
screen "MTA-ChillersBombasEnvasado" 800x480, template "Plantilla_2"
   GraphicView "Visor de gráficos_3" at 648,158 size 48x71; Picture "Bomba"
   GraphicIOField "Plantilla_Campo ES gráfico_2" at 684,217 size 49x36; PictureList "Motor2"
      ProcessValue <- "AnimaciónMT009"
   SymbolicIOField "Campo ES simbólico_4" at 602,132 size 172x21; TextOff '0'; TextOn '1'; TextList "EstadoMotor"
      ProcessValue <- "AnimaciónMT009"
   TextField "Campo de texto_6" at 599,93 size 42x18; Text 'MT009'
   GraphicView "Visor de gráficos_4" at 454,158 size 48x71; Picture "Bomba"
   GraphicIOField "Plantilla_Campo ES gráfico_1" at 490,217 size 49x36; PictureList "Motor2"
      ProcessValue <- "AnimaciónMT010"
   SymbolicIOField "Campo ES simbólico_1" at 408,132 size 172x21; TextOff '0'; TextOn '1'; TextList "EstadoMotor"
      ProcessValue <- "AnimaciónMT010"
   TextField "Campo de texto_7" at 405,93 size 42x18; Text 'MT010'
   GraphicView "Visor de gráficos_6" at 64,158 size 48x71; Picture "Bomba"
   GraphicIOField "Plantilla_Campo ES gráfico_4" at 100,217 size 49x36; PictureList "Motor2"
      ProcessValue <- "AnimaciónMP013"
   SymbolicIOField "Campo ES simbólico_3" at 20,132 size 172x21; TextOff '0'; TextOn '1'; TextList "EstadoMotor"
      ProcessValue <- "AnimaciónMP013"
   TextField "Campo de texto_9" at 23,93 size 41x18; Text 'MP013'
   TextField "Campo de texto_19" at 405,112 size 169x18; Text 'Intercambiador Línea 1 y Man.'
   GraphicView "Visor de gráficos_5" at 260,158 size 48x71; Picture "Bomba"
   GraphicIOField "Plantilla_Campo ES gráfico_3" at 296,217 size 49x36; PictureList "Motor2"
      ProcessValue <- "AnimaciónMP012"
   SymbolicIOField "Campo ES simbólico_2" at 214,132 size 172x21; TextOff '0'; TextOn '1'; TextList "EstadoMotor"
      ProcessValue <- "AnimaciónMP012"
   TextField "Campo de texto_8" at 211,93 size 41x18; Text 'MP012'
   TextField "Campo de texto_18" at 598,112 size 150x18; Text 'Intercambiador Línea 3 y 5'
   TextField "Campo de texto_16" at 215,113 size 150x18; Text 'Chillers Envasado - Principal'
   TextField "Campo de texto_17" at 21,113 size 146x18; Text 'Chillers Envasado - Backup'
   GraphicView "Plantilla_Visor de gráficos_2" at 752,6 size 35x35; Picture "ParlantesGris_1"
   GraphicView "Plantilla_Visor de gráficos_1" at 752,6 size 35x35; Picture "ParlantesRojo"
      Visibility <- "SirenaChillers"
   Button "Botón_1" at 740,1 size 57x44; TextOff 'Text'
      on Click: ActivateScreen("MTA-ChillersConfiguraciónSirena", 0)
   ScreenModuleView "ControlMotor-NoAUTO_1" at 609,271 size 163x76
      Guid_{11997190-67152} <- "DesMT009"
      Guid_{11997190-67156} <- "ParadaMT009"
      Guid_{11997190-67150} <- "HabMT009"
      Guid_{11997190-67154} <- "MarchaMT009"
   ScreenModuleView "ControlMotor-NoAUTO_2" at 413,271 size 163x76
      Guid_{11997190-67152} <- "DesMT010"
      Guid_{11997190-67156} <- "ParadaMT010"
      Guid_{11997190-67150} <- "HabMT010"
      Guid_{11997190-67154} <- "MarchaMT010"
   ScreenModuleView "ControlMotor-NoAUTO_3" at 219,271 size 163x76
      Guid_{11997190-67152} <- "DesMP012"
      Guid_{11997190-67156} <- "ParadaMP012"
      Guid_{11997190-67150} <- "HabMP012"
      Guid_{11997190-67154} <- "MarchaMP012"
   ScreenModuleView "ControlMotor-NoAUTO_4" at 22,271 size 163x76
      Guid_{11997190-67152} <- "DesMP013"
      Guid_{11997190-67156} <- "ParadaMP013"
      Guid_{11997190-67150} <- "HabMP013"
      Guid_{11997190-67154} <- "MarchaMP013"
   TextField "Campo de texto_5" at 256,10 size 261x27; Text 'Chillers - Bombas de Envasado'

screen "MTA-ChillersBombasSoplado" 800x480, template "Plantilla_2"
   TextField "Campo de texto_5" at 256,10 size 248x27; Text 'Chillers - Bombas de Soplado'
   GraphicView "Visor de gráficos_3" at 648,158 size 48x71; Picture "Bomba"
   GraphicIOField "Plantilla_Campo ES gráfico_8" at 684,217 size 49x36; PictureList "Motor2"
      ProcessValue <- "AnimaciónMT007"
   SymbolicIOField "Campo ES simbólico_4" at 602,132 size 172x21; TextOff '0'; TextOn '1'; TextList "EstadoMotor"
      ProcessValue <- "AnimaciónMT007"
   TextField "Campo de texto_6" at 599,93 size 42x18; Text 'MT007'
   GraphicView "Visor de gráficos_4" at 454,158 size 48x71; Picture "Bomba"
   GraphicIOField "Plantilla_Campo ES gráfico_7" at 490,217 size 49x36; PictureList "Motor2"
      ProcessValue <- "AnimaciónMT008"
   SymbolicIOField "Campo ES simbólico_1" at 408,132 size 172x21; TextOff '0'; TextOn '1'; TextList "EstadoMotor"
      ProcessValue <- "AnimaciónMT008"
   TextField "Campo de texto_7" at 405,93 size 42x18; Text 'MT008'
   GraphicView "Visor de gráficos_6" at 64,158 size 48x71; Picture "Bomba"
   GraphicIOField "Plantilla_Campo ES gráfico_5" at 100,217 size 49x36; PictureList "Motor2"
      ProcessValue <- "AnimaciónMP011"
   SymbolicIOField "Campo ES simbólico_3" at 20,132 size 172x21; TextOff '0'; TextOn '1'; TextList "EstadoMotor"
      ProcessValue <- "AnimaciónMP011"
   TextField "Campo de texto_9" at 23,93 size 41x18; Text 'MP011'
   TextField "Campo de texto_19" at 407,113 size 140x18; Text 'Sopladora Línea 3 y Man.'
   GraphicView "Visor de gráficos_5" at 260,158 size 48x71; Picture "Bomba"
   GraphicIOField "Plantilla_Campo ES gráfico_6" at 296,217 size 49x36; PictureList "Motor2"
      ProcessValue <- "AnimaciónMP010"
   SymbolicIOField "Campo ES simbólico_2" at 214,132 size 172x21; TextOff '0'; TextOn '1'; TextList "EstadoMotor"
      ProcessValue <- "AnimaciónMP010"
   TextField "Campo de texto_8" at 211,93 size 41x18; Text 'MP010'
   TextField "Campo de texto_18" at 599,113 size 104x18; Text 'Sopladora Línea 1'
   TextField "Campo de texto_16" at 212,113 size 142x18; Text 'Chillers Soplado - Principal'
   TextField "Campo de texto_17" at 21,113 size 138x18; Text 'Chillers Soplado - Backup'
   GraphicView "Plantilla_Visor de gráficos_2" at 752,6 size 35x35; Picture "ParlantesGris_1"
   GraphicView "Plantilla_Visor de gráficos_1" at 752,6 size 35x35; Picture "ParlantesRojo"
      Visibility <- "SirenaChillers"
   Button "Botón_1" at 740,1 size 57x44; TextOff 'Text'
      on Click: ActivateScreen("MTA-ChillersConfiguraciónSirena", 0)
   ScreenModuleView "ControlMotor-NoAUTO_1" at 609,271 size 163x76
      Guid_{11997190-67152} <- "DesMT007"
      Guid_{11997190-67156} <- "ParadaMT007"
      Guid_{11997190-67150} <- "HabMT007"
      Guid_{11997190-67154} <- "MarchaMT007"
   ScreenModuleView "ControlMotor-NoAUTO_3" at 219,271 size 163x76
      Guid_{11997190-67152} <- "DesMP010"
      Guid_{11997190-67156} <- "ParadaMP010"
      Guid_{11997190-67150} <- "HabMP010"
      Guid_{11997190-67154} <- "MarchaMP010"
   ScreenModuleView "ControlMotor-NoAUTO_2" at 417,271 size 163x76
      Guid_{11997190-67152} <- "DesMT008"
      Guid_{11997190-67156} <- "ParadaMT008"
      Guid_{11997190-67150} <- "HabMT008"
      Guid_{11997190-67154} <- "MarchaMT008"
   ScreenModuleView "ControlMotor-NoAUTO_4" at 27,271 size 163x76
      Guid_{11997190-67152} <- "DesMP011"
      Guid_{11997190-67156} <- "ParadaMP011"
      Guid_{11997190-67150} <- "HabMP011"
      Guid_{11997190-67154} <- "MarchaMP011"

screen "MTA-ChillersConfiguraciónSirena" 800x480, template "Plantilla_2"
   Switch "Interruptor_1" at 119,81 size 36x32; TextOn 'Habilitado'; CaptionText 'Switch'; TextOff 'Deshabilitado'; PictureOff "ParlantesGrisClaro_1"; PictureOn "ParlantesVerde2_1"
      ProcessValue <- "SirenaM1"
   Switch "Interruptor_2" at 119,118 size 36x32; TextOn 'Habilitado'; CaptionText 'Switch'; TextOff 'Deshabilitado'; PictureOff "ParlantesGrisClaro_1"; PictureOn "ParlantesVerde2_1"
      ProcessValue <- "SirenaM2"
   Switch "Interruptor_3" at 119,155 size 36x32; TextOn 'Habilitado'; CaptionText 'Switch'; TextOff 'Deshabilitado'; PictureOff "ParlantesGrisClaro_1"; PictureOn "ParlantesVerde2_1"
      ProcessValue <- "SirenaM3"
   Switch "Interruptor_4" at 119,192 size 36x32; TextOn 'Habilitado'; CaptionText 'Switch'; TextOff 'Deshabilitado'; PictureOff "ParlantesGrisClaro_1"; PictureOn "ParlantesVerde2_1"
      ProcessValue <- "SirenaM4"
   Switch "Interruptor_5" at 119,229 size 36x32; TextOn 'Habilitado'; CaptionText 'Switch'; TextOff 'Deshabilitado'; PictureOff "ParlantesGrisClaro_1"; PictureOn "ParlantesVerde2_1"
      ProcessValue <- "SirenaM5"
   TextField "Campo de texto_1" at 163,233 size 365x22; Text 'Ninguna Bomba para torres de enfriamiento en marcha'
   TextField "Campo de texto_2" at 163,196 size 424x22; Text 'Ninguna Bomba para Intercambiadores de Envasado en marcha'
   TextField "Campo de texto_3" at 163,160 size 353x22; Text 'Ninguna Bomba para Chillers de Envasado en marcha'
   TextField "Campo de texto_4" at 163,122 size 411x22; Text 'Ninguna Bomba para Intercambiadores de Solpado en marcha'
   TextField "Campo de texto_5" at 163,86 size 340x22; Text 'Ninguna Bomba para Chillers de Soplado en marcha'
   TextField "Campo de texto_6" at 51,53 size 277x22; Text 'Motivos para que la sirena se active:'
   TextField "Campo de texto_7" at 214,8 size 319x29; Text 'Chillers - Configuración de Sirena'
   Switch "Interruptor_6" at 119,266 size 36x32; TextOn 'Habilitado'; CaptionText 'Switch'; TextOff 'Deshabilitado'; PictureOff "ParlantesGrisClaro_1"; PictureOn "ParlantesVerde2_1"
      ProcessValue <- "SirenaM6"
   TextField "Campo de texto_8" at 163,271 size 231x22; Text 'Ningún Chiller de Soplado Habilitado'
   Switch "Interruptor_7" at 119,303 size 36x32; TextOn 'Habilitado'; CaptionText 'Switch'; TextOff 'Deshabilitado'; PictureOff "ParlantesGrisClaro_1"; PictureOn "ParlantesVerde2_1"
      ProcessValue <- "SirenaM7"
   TextField "Campo de texto_9" at 163,307 size 244x22; Text 'Ningún Chiller de Envasado Habilitado'
   Switch "Interruptor_8" at 119,341 size 36x32; TextOn 'Habilitado'; CaptionText 'Switch'; TextOff 'Deshabilitado'; PictureOff "ParlantesGrisClaro_1"; PictureOn "ParlantesVerde2_1"
      ProcessValue <- "SirenaM8"
   TextField "Campo de texto_10" at 163,346 size 150x22; Text 'Alarma en algún Chiller'
   GraphicView "Plantilla_Visor de gráficos_2" at 752,6 size 35x35; Picture "ParlantesGris_1"
   GraphicView "Plantilla_Visor de gráficos_1" at 752,6 size 35x35; Picture "ParlantesRojo"
      Visibility <- "SirenaChillers"
   Button "Botón_1" at 740,1 size 57x44; TextOff 'Text'
      on Click: ActivateScreen("MTA-ChillersConfiguraciónSirena", 0)
   Switch "Interruptor_9" at 119,378 size 36x32; TextOn 'Habilitado'; CaptionText 'Switch'; TextOff 'Deshabilitado'; PictureOff "ParlantesGrisClaro_1"; PictureOn "ParlantesVerde2_1"
      ProcessValue <- "SirenaM9"
   TextField "Campo de texto_11" at 163,383 size 194x22; Text 'Falla Térmica en algún motor'

screen "MTA-Chillers-Envasado" 800x480, template "Plantilla_2"
   GraphicView "Visor de gráficos_2" at 24,127 size 192x232; Picture "Chiller2b"
   GraphicView "Visor de gráficos_1" at 432,129 size 144x104; Picture "Chillerb"
   Switch "Interruptor_1" at 243,127 size 91x31; TextOff 'Habilitado'; TextOn 'Deshabilitado'; CaptionText 'Switch'
      Appearance <- "Habilitación-CH-ENV-GR"
      ProcessValue <- "Habilitación-CH-ENV-GR"
   TextField "Campo de texto_5" at 309,10 size 182x27; Text 'Chillers de Envasado'
   TextField "Campo de texto_10" at 19,78 size 169x22; Text 'Chiller Envasado GRANDE'
   TextField "Campo de texto_6" at 411,78 size 158x22; Text 'Chiller Envasado CHICO'
   Circle "Círculo_9" at 243,225 size 16x16
      Appearance <- "MAX-CH-ENV-GR"
   Circle "Círculo_10" at 243,183 size 16x16
      Appearance <- "RUN-CH-ENV-GR"
   Circle "Círculo_11" at 243,204 size 16x16
      Appearance <- "Alarma1-CH-ENV-GR"
   TextField "Campo de texto_1" at 263,203 size 40x18; Text 'Alarma'
   TextField "Campo de texto_3" at 263,182 size 108x18; Text 'En Funcionamiento'
   TextField "Campo de texto_4" at 263,223 size 101x18; Text 'Máxima Capacidad'
   Switch "Interruptor_2" at 595,127 size 91x31; TextOff 'Habilitado'; TextOn 'Deshabilitado'; CaptionText 'Switch'
      Appearance <- "Habilitación-CH-ENV-CH"
      ProcessValue <- "Habilitación-CH-ENV-CH"
   GraphicView "Plantilla_Visor de gráficos_2" at 752,6 size 35x35; Picture "ParlantesGris_1"
   GraphicView "Plantilla_Visor de gráficos_1" at 752,6 size 35x35; Picture "ParlantesRojo"
      Visibility <- "SirenaChillers"
   Button "Botón_1" at 740,1 size 57x44; TextOff 'Text'
      on Click: ActivateScreen("MTA-ChillersConfiguraciónSirena", 0)
   TextField "Campo de texto_24" at 613,183 size 79x18; Text 'Alarma Aceite'
   TextField "Campo de texto_25" at 613,166 size 108x18; Text 'En Funcionamiento'
   TextField "Campo de texto_26" at 613,201 size 115x18; Text 'Alarma Temperatura'
   TextField "Campo de texto_27" at 613,220 size 125x18; Text 'Alarma Térmico motor'
   Circle "Círculo_2" at 593,167 size 16x16
      Appearance <- "CH-ENV-CH-RUN"
   Circle "Círculo_3" at 593,185 size 16x16
      Appearance <- "CH-ENV-CH-ACT"
   Circle "Círculo_5" at 593,204 size 16x16
      Appearance <- "CH-ENV-CH-TEMP"
   Circle "Círculo_6" at 593,223 size 16x16
      Appearance <- "CH-ENV-CH-TERM"

screen "MTA-Chillers-General" 800x480, template "Plantilla_2"
   GraphicView "Visor de gráficos_7" at 488,183 size 48x71; Picture "Bomba"
   GraphicView "Visor de gráficos_8" at 536,183 size 48x71; Picture "Bomba"
   GraphicView "Visor de gráficos_1" at 392,183 size 48x71; Picture "Bomba"
   GraphicView "Visor de gráficos_9" at 440,183 size 48x71; Picture "Bomba"
   GraphicView "Visor de gráficos_17" at 383,130 size 87x77; Picture "tubo"
   GraphicView "Visor de gráficos_18" at 479,130 size 87x77; Picture "tubo"
   GraphicView "Visor de gráficos_14" at 384,48 size 141x131; Picture "Tanque3_1"
   GraphicView "Visor de gráficos_3" at 750,189 size 48x212; Picture "Chiller2bb"
   GraphicView "Visor de gráficos_4" at 630,161 size 96x96; Picture "Chiller_2"
   GraphicView "Visor de gráficos_5" at 264,183 size 48x71; Picture "Bomba"
   GraphicView "Visor de gráficos_6" at 312,183 size 48x71; Picture "Bomba"
   GraphicView "Visor de gráficos_10" at 168,183 size 48x71; Picture "Bomba"
   GraphicView "Visor de gráficos_11" at 216,183 size 48x71; Picture "Bomba"
   GraphicView "Visor de gráficos_2" at 12,132 size 128x144; Picture "Chiller2b"
   GraphicView "Visor de gráficos_12" at 45,333 size 88x77; Picture "Chillerb"
   GraphicView "Visor de gráficos_15" at 159,130 size 87x77; Picture "tubo"
   GraphicView "Visor de gráficos_16" at 255,130 size 87x77; Picture "tubo"
   GraphicView "Visor de gráficos_13" at 162,48 size 141x131; Picture "Tanque3_1"
   GraphicIOField "Plantilla_Campo ES gráfico_2" at 304,240 size 41x36; PictureList "Motor2"
      ProcessValue <- "AnimaciónMT010"
   GraphicIOField "Plantilla_Campo ES gráfico_1" at 352,240 size 41x36; PictureList "Motor2"
      ProcessValue <- "AnimaciónMT009"
   GraphicIOField "Plantilla_Campo ES gráfico_3" at 528,240 size 41x36; PictureList "Motor2"
      ProcessValue <- "AnimaciónMT008"
   GraphicIOField "Plantilla_Campo ES gráfico_4" at 576,240 size 41x36; PictureList "Motor2"
      ProcessValue <- "AnimaciónMT007"
   GraphicIOField "Plantilla_Campo ES gráfico_5" at 432,240 size 41x36; PictureList "Motor2"
      ProcessValue <- "AnimaciónMP011"
   GraphicIOField "Plantilla_Campo ES gráfico_6" at 480,240 size 41x36; PictureList "Motor2"
      ProcessValue <- "AnimaciónMP010"
   GraphicIOField "Plantilla_Campo ES gráfico_7" at 208,240 size 41x36; PictureList "Motor2"
      ProcessValue <- "AnimaciónMP013"
   GraphicIOField "Plantilla_Campo ES gráfico_8" at 256,240 size 41x36; PictureList "Motor2"
      ProcessValue <- "AnimaciónMP012"
   TextField "Campo de texto_1" at 631,124 size 86x32; Text 'Chiller Soplado Chico'
   TextField "Campo de texto_2" at 668,364 size 86x32; Text 'Chiller Soplado Grande'
   TextField "Campo de texto_3" at 142,373 size 90x32; Text 'Chiller Envasado Chico'
   TextField "Campo de texto_4" at 28,94 size 90x32; Text 'Chiller Envasado Grande'
   TextField "Campo de texto_5" at 334,8 size 72x29; Text 'Chillers'
   TextField "Campo de texto_6" at 474,309 size 131x25; Text 'Bombas Soplado'
   TextField "Campo de texto_7" at 242,309 size 139x25; Text 'Bombas Envasado'
   TextField "Campo de texto_9" at 520,70 size 51x52; Text 'Tanque Soplado'
   TextField "Campo de texto_8" at 214,277 size 41x19; Text 'MP013'
   TextField "Campo de texto_11" at 262,277 size 41x19; Text 'MP012'
   TextField "Campo de texto_12" at 310,277 size 49x19; Text 'MT010'
   TextField "Campo de texto_13" at 366,277 size 42x19; Text 'MT009'
   TextField "Campo de texto_14" at 438,277 size 41x19; Text 'MP011'
   TextField "Campo de texto_15" at 486,277 size 41x19; Text 'MP010'
   TextField "Campo de texto_16" at 534,277 size 42x19; Text 'MT008'
   TextField "Campo de texto_17" at 590,277 size 42x19; Text 'MT007'
   TextField "Campo de texto_10" at 294,69 size 58x52; Text 'Tanque Envasado'
   Button "Botón_3" at 629,155 size 170x254; TextOff 'Control Soplado'
      on Click: ActivateScreen("MTA-Chillers-Soplado", 0)
   Button "Botón_2" at 419,227 size 215x78; TextOff 'Control Soplado'
      on Click: ActivateScreen("MTA-ChillersBombasSoplado", 0)
   Button "Botón_4" at 0,122 size 194x294; TextOff 'Control Soplado'
      on Click: ActivateScreen("MTA-Chillers-Envasado", 0)
   Button "Botón_5" at 203,226 size 208x79; TextOff 'Control Envasado'
      on Click: ActivateScreen("MTA-ChillersBombasEnvasado", 0)
   Circle "Círculo_5" at 722,327 size 16x16
      Appearance <- "MAX-CH-SOP-GR"
   Circle "Círculo_6" at 722,292 size 16x16
      Appearance <- "RUN-CH-SOP-GR"
   Circle "Círculo_8" at 722,310 size 16x16
      Appearance <- "Alarma1-CH-SOP-GR"
   Circle "Círculo_1" at 147,255 size 16x16
      Appearance <- "MAX-CH-ENV-GR"
   Circle "Círculo_2" at 147,220 size 16x16
      Appearance <- "RUN-CH-ENV-GR"
   Circle "Círculo_3" at 147,238 size 16x16
      Appearance <- "Alarma1-CH-ENV-GR"
   Circle "Círculo_4" at 18,338 size 16x16
      Appearance <- "RUN-CH-ENV-CH"
   GraphicView "Plantilla_Visor de gráficos_2" at 752,6 size 35x35; Picture "ParlantesGris_1"
   GraphicView "Plantilla_Visor de gráficos_1" at 752,6 size 35x35; Picture "ParlantesRojo"
      Visibility <- "SirenaChillers"
   Button "Botón_1" at 740,1 size 57x44; TextOff 'Text'
      on Click: ActivateScreen("MTA-ChillersConfiguraciónSirena", 0)
   Circle "Círculo_7" at 18,355 size 16x16
      Appearance <- "CH-ENV-CH-ACT"
   Circle "Círculo_9" at 18,372 size 16x16
      Appearance <- "CH-ENV-CH-TEMP"
   Circle "Círculo_10" at 18,389 size 16x16
      Appearance <- "CH-ENV-CH-TERM"
   Circle "Círculo_11" at 606,165 size 16x16
      Appearance <- "CH-SOP-CH-CTC1ON"
   Circle "Círculo_12" at 606,182 size 16x16
      Appearance <- "CH-SOP-CH-CTC2ON"
   Circle "Círculo_14" at 606,217 size 16x16
      Appearance <- "CH-SOP-CH-TERM1"

screen "MTA-Chillers-Soplado" 800x480, template "Plantilla_2"
   GraphicView "Visor de gráficos_2" at 24,127 size 192x232; Picture "Chiller2c"
   GraphicView "Visor de gráficos_1" at 424,129 size 160x168; Picture "Chiller_2"
   Switch "Interruptor_1" at 243,127 size 91x31; TextOff 'Habilitado'; TextOn 'Deshabilitado'; CaptionText 'Switch'
      Appearance <- "Habilitación-CH-SOP-GR"
      ProcessValue <- "Habilitación-CH-SOP-GR"
   TextField "Campo de texto_1" at 263,203 size 40x18; Text 'Alarma'
   TextField "Campo de texto_3" at 263,182 size 108x18; Text 'En Funcionamiento'
   TextField "Campo de texto_4" at 263,223 size 101x18; Text 'Máxima Capacidad'
   TextField "Campo de texto_5" at 311,10 size 169x27; Text 'Chillers de Soplado'
   TextField "Campo de texto_10" at 19,78 size 156x22; Text 'Chiller Soplado GRANDE'
   TextField "Campo de texto_6" at 411,78 size 145x22; Text 'Chiller Soplado CHICO'
   Circle "Círculo_5" at 242,225 size 16x16
      Appearance <- "MAX-CH-SOP-GR"
   Circle "Círculo_6" at 242,182 size 16x16
      Appearance <- "RUN-CH-SOP-GR"
   Circle "Círculo_8" at 242,204 size 16x16
      Appearance <- "Alarma1-CH-SOP-GR"
   Switch "Interruptor_2" at 627,127 size 91x31; TextOff 'Habilitado'; TextOn 'Deshabilitado'; CaptionText 'Switch'
      Appearance <- "Habilitación-CH-SOP-CH"
      ProcessValue <- "Habilitación-CH-SOP-CH"
   GraphicView "Plantilla_Visor de gráficos_2" at 752,6 size 35x35; Picture "ParlantesGris_1"
   GraphicView "Plantilla_Visor de gráficos_1" at 752,6 size 35x35; Picture "ParlantesRojo"
      Visibility <- "SirenaChillers"
   Button "Botón_1" at 740,1 size 57x44; TextOff 'Text'
      on Click: ActivateScreen("MTA-ChillersConfiguraciónSirena", 0)
   TextField "Campo de texto_28" at 607,198 size 120x18; Text 'Motor 2 Funcionando'
   TextField "Campo de texto_29" at 607,177 size 120x18; Text 'Motor 1 Funcionando'
   TextField "Campo de texto_30" at 631,220 size 96x18; Text 'Térmico motor 1'
   TextField "Campo de texto_31" at 631,241 size 96x18; Text 'Térmico motor 2'
   Circle "Círculo_11" at 734,181 size 16x16
      Appearance <- "CH-SOP-CH-CTC1ON"
   Circle "Círculo_12" at 734,200 size 16x16
      Appearance <- "CH-SOP-CH-CTC2ON"
   Circle "Círculo_14" at 734,240 size 16x16
      Appearance <- "CH-SOP-CH-TERM1"

screen "MTA-TorreEnfriamientoBMB" 800x480, template "Plantilla_2"
   GraphicView "Visor de gráficos_1" at 167,153 size 98x119; Picture "torreFINAL4_1"
   GraphicView "Visor de gráficos_4" at 260,143 size 138x153; Picture "torreFINAL4_1"
   GraphicView "Visor de gráficos_17" at 16,128 size 178x201; Picture "torreFINAL4_1"
   GraphicView "Visor de gráficos_2" at 167,153 size 98x119; Picture "torreFINAL4B_1"
   GraphicView "Visor de gráficos_3" at 260,143 size 138x153; Picture "torreFINAL4B_1"
   GraphicView "Visor de gráficos_5" at 16,128 size 178x201; Picture "torreFINAL4B_1"
   GraphicView "Visor de gráficos_6" at 167,153 size 98x119; Picture "torreFINAL4C_1"
      Visibility <- "BombaTorreON"
   GraphicView "Visor de gráficos_15" at 260,143 size 138x153; Picture "torreFINAL4C_1"
      Visibility <- "BombaTorreON"
   GraphicView "Visor de gráficos_16" at 16,128 size 178x201; Picture "torreFINAL4C_1"
      Visibility <- "BombaTorreON"
   TextField "Campo de texto_1" at 361,84 size 57x23; Text 'Torre 2'
   TextField "Campo de texto_2" at 229,95 size 47x20; Text 'Torre 3'
   TextField "Campo de texto_12" at 101,76 size 57x23; Text 'Torre 1'
   TextField "Campo de texto_13" at 273,197 size 55x29; Text 'Norte'
   TextField "Campo de texto_14" at 38,202 size 50x34; Text 'Este'
   GraphicIOField "Campo ES gráfico_1" at 76,122 size 56x29; PictureList "MotorTorre"
      ProcessValue <- "AnimaciónV001"
   GraphicIOField "Campo ES gráfico_2" at 199,147 size 33x21; PictureList "MotorTorre"
      ProcessValue <- "AnimaciónV003"
   GraphicIOField "Campo ES gráfico_3" at 306,137 size 45x24; PictureList "MotorTorre"
      ProcessValue <- "AnimaciónV002"
   GraphicView "Visor de gráficos_19" at 0,384 size 800x15; Picture "TUBOXXX"
   GraphicView "Plantilla_Visor de gráficos_2" at 752,6 size 35x35; Picture "ParlantesGris_1"
   GraphicView "Plantilla_Visor de gráficos_1" at 752,6 size 35x35; Picture "ParlantesRojo"
      Visibility <- "SirenaChillers"
   Button "Botón_1" at 740,1 size 57x44; TextOff 'Text'
      on Click: ActivateScreen("MTA-ChillersConfiguraciónSirena", 0)
   Button "Botón_2" at 200,320 size 152x38; TextOff 'VENTILADORES'
      on Click: ActivateScreen("MTA-TorreEnfriamientoVENT", 0)
   TextField "Campo de texto_10" at 41,374 size 98x32; Text 'Presostato Agua Torres'
   TextField "Campo de texto_5" at 238,8 size 293x29; Text 'Torres de enfriamiento Chillers'
   GraphicView "Visor de gráficos_9" at 30,56 size 63x62; Picture "Vent1"
   GraphicView "Visor de gráficos_10" at 30,56 size 63x62; Picture "Vent2"
      Visibility <- "AnimaciónV001"
   GraphicView "Visor de gráficos_11" at 177,82 size 47x46; Picture "Vent1"
   GraphicView "Visor de gráficos_12" at 177,82 size 47x46; Picture "Vent2"
      Visibility <- "AnimaciónV003"
   GraphicView "Visor de gráficos_13" at 292,66 size 63x62; Picture "Vent1"
   GraphicView "Visor de gráficos_14" at 292,66 size 63x62; Picture "Vent2"
      Visibility <- "AnimaciónV002"
   IOField "Campo ES_1" at 241,360 size 80x23; FormatPattern 999.99; Unit  ºC
      ProcessValue <- "TemperaturatorresCH"
   GraphicView "Visor de gráficos_8" at 459,277 size 48x71; Picture "Bomba"
   GraphicIOField "Plantilla_Campo ES gráfico_1" at 497,336 size 49x36; PictureList "Motor2"
      ProcessValue <- "AnimaciónMP019"
   SymbolicIOField "Campo ES simbólico_1" at 581,259 size 172x20; TextOff '0'; TextOn '1'; TextList "EstadoMotor"
      ProcessValue <- "AnimaciónMP019"
   TextField "Campo de texto_7" at 495,293 size 41x18; Text 'MP019'
   TextField "Campo de texto_17" at 455,241 size 129x27; Text 'Backup (ESTE)'
   ScreenModuleView "ControlMotor-NoAUTO_4" at 565,285 size 203x76
      Guid_{11997190-67152} <- "DesMP019"
      Guid_{11997190-67156} <- "ParadaMP019"
      Guid_{11997190-67150} <- "HabMP019"
      Guid_{11997190-67154} <- "MarchaMP019"
   ScreenModuleView "ControlMotor-NoAUTO_1" at 564,115 size 203x76
      Guid_{11997190-67152} <- "DesMP018"
      Guid_{11997190-67156} <- "ParadaMP018"
      Guid_{11997190-67150} <- "HabMP018"
      Guid_{11997190-67154} <- "MarchaMP018"
   SymbolicIOField "Campo ES simbólico_4" at 575,89 size 172x20; TextOff '0'; TextOn '1'; TextList "EstadoMotor"
      ProcessValue <- "AnimaciónMP018"
   TextField "Campo de texto_6" at 494,129 size 41x18; Text 'MP018'
   TextField "Campo de texto_16" at 454,77 size 151x27; Text 'Principal (OESTE)'
   GraphicView "Visor de gráficos_7" at 458,113 size 48x71; Picture "Bomba"
   GraphicIOField "Plantilla_Campo ES gráfico_2" at 496,172 size 49x36; PictureList "Motor2"
      ProcessValue <- "AnimaciónMP018"

screen "MTA-TorreEnfriamientoVENT" 800x480, template "Plantilla_2"
   GraphicView "Visor de gráficos_1" at 167,153 size 98x119; Picture "torreFINAL4_1"
   GraphicView "Visor de gráficos_4" at 260,143 size 138x153; Picture "torreFINAL4_1"
   GraphicView "Visor de gráficos_17" at 16,128 size 178x201; Picture "torreFINAL4_1"
   GraphicView "Visor de gráficos_2" at 167,153 size 98x119; Picture "torreFINAL4B_1"
   GraphicView "Visor de gráficos_3" at 260,143 size 138x153; Picture "torreFINAL4B_1"
   GraphicView "Visor de gráficos_5" at 16,128 size 178x201; Picture "torreFINAL4B_1"
   GraphicView "Visor de gráficos_6" at 167,153 size 98x119; Picture "torreFINAL4C_1"
      Visibility <- "BombaTorreON"
   GraphicView "Visor de gráficos_15" at 260,143 size 138x153; Picture "torreFINAL4C_1"
      Visibility <- "BombaTorreON"
   GraphicView "Visor de gráficos_16" at 16,128 size 178x201; Picture "torreFINAL4C_1"
      Visibility <- "BombaTorreON"
   SymbolicIOField "Campo ES simbólico_2" at 548,59 size 188x19; TextOff '0'; TextOn '1'; TextList "EstadoMotor"
      ProcessValue <- "AnimaciónV001"
   SymbolicIOField "Campo ES simbólico_3" at 549,181 size 188x19; TextOff '0'; TextOn '1'; TextList "EstadoMotor"
      ProcessValue <- "AnimaciónV002"
   SymbolicIOField "Campo ES simbólico_7" at 549,301 size 188x19; TextOff '0'; TextOn '1'; TextList "EstadoMotor"
      ProcessValue <- "AnimaciónV003"
   TextField "Campo de texto_1" at 361,84 size 57x23; Text 'Torre 2'
   TextField "Campo de texto_2" at 229,95 size 47x20; Text 'Torre 3'
   TextField "Campo de texto_13" at 273,197 size 55x29; Text 'Norte'
   TextField "Campo de texto_14" at 38,202 size 50x34; Text 'Este'
   ScreenModuleView "Faceplate_4_1" at 447,84 size 245x68
      Guid_{11997190-23979} <- "HabV001(1)"
      Guid_{11997190-23983} <- "ParadaV001(1)"
      Guid_{11997190-23981} <- "MarchaV001(1)"
      Guid_{11997190-23989} <- "SP-OFF-V001"
      Guid_{11997190-23976} <- "DeshV001"
      Guid_{11997190-23987} <- "SP-ON-V001"
      Guid_{11997190-23985} <- "AnimaMenuV001"
   TextField "Campo de texto_4" at 439,176 size 104x27; Text 'Ventilador 2'
   TextField "Campo de texto_3" at 439,54 size 104x27; Text 'Ventilador 1'
   TextField "Campo de texto_23" at 440,298 size 104x27; Text 'Ventilador 3'
   ScreenModuleView "Faceplate_4_2" at 447,204 size 245x68
      Guid_{11997190-23979} <- "HabV002(1)"
      Guid_{11997190-23983} <- "ParadaV002(1)"
      Guid_{11997190-23981} <- "MarchaV002(1)"
      Guid_{11997190-23989} <- "SP-OFF-V002"
      Guid_{11997190-23976} <- "DeshV002"
      Guid_{11997190-23987} <- "SP-ON-V002"
      Guid_{11997190-23985} <- "AnimaMenuV002"
   ScreenModuleView "Faceplate_4_3" at 447,326 size 245x68
      Guid_{11997190-23979} <- "HabV003(1)"
      Guid_{11997190-23983} <- "ParadaV003(1)"
      Guid_{11997190-23981} <- "MarchaV003(1)"
      Guid_{11997190-23989} <- "SP-OFF-V003"
      Guid_{11997190-23976} <- "DeshV003"
      Guid_{11997190-23987} <- "SP-ON-V003"
      Guid_{11997190-23985} <- "AnimaMenuV003"
   TextField "Campo de texto_12" at 101,76 size 57x23; Text 'Torre 1'
   GraphicIOField "Campo ES gráfico_1" at 76,122 size 56x29; PictureList "MotorTorre"
      ProcessValue <- "AnimaciónV001"
   GraphicIOField "Campo ES gráfico_2" at 199,147 size 33x21; PictureList "MotorTorre"
      ProcessValue <- "AnimaciónV003"
   GraphicIOField "Campo ES gráfico_3" at 306,137 size 45x24; PictureList "MotorTorre"
      ProcessValue <- "AnimaciónV002"
   Switch "Interruptor_1" at 744,62 size 32x29; TextOn 'Auto'; CaptionText 'Switch'; TextOff 'Manual'; PictureOff "A2"; PictureOn "A"
      Appearance <- "AutoV001"
      ProcessValue <- "AutoV001"
   Switch "Interruptor_2" at 744,184 size 32x29; TextOn 'Auto'; CaptionText 'Switch'; TextOff 'Manual'; PictureOff "A2"; PictureOn "A"
      Appearance <- "AutoV002"
      ProcessValue <- "AutoV002"
   Switch "Interruptor_3" at 744,304 size 32x29; TextOn 'Auto'; CaptionText 'Switch'; TextOff 'Manual'; PictureOff "A2"; PictureOn "A"
      Appearance <- "AutoV003"
      ProcessValue <- "AutoV003"
   GraphicView "Visor de gráficos_19" at 0,384 size 800x15; Picture "TUBOXXX"
   TextField "Campo de texto_5" at 238,8 size 293x29; Text 'Torres de enfriamiento Chillers'
   GraphicView "Visor de gráficos_9" at 30,56 size 63x62; Picture "Vent1"
   GraphicView "Visor de gráficos_10" at 30,56 size 63x62; Picture "Vent2"
      Visibility <- "AnimaciónV001"
   GraphicView "Visor de gráficos_11" at 177,82 size 47x46; Picture "Vent1"
   GraphicView "Visor de gráficos_12" at 177,82 size 47x46; Picture "Vent2"
      Visibility <- "AnimaciónV003"
   GraphicView "Visor de gráficos_13" at 292,66 size 63x62; Picture "Vent1"
   GraphicView "Visor de gráficos_14" at 292,66 size 63x62; Picture "Vent2"
      Visibility <- "AnimaciónV002"
   GraphicView "Plantilla_Visor de gráficos_2" at 752,6 size 35x35; Picture "ParlantesGris_1"
   GraphicView "Plantilla_Visor de gráficos_1" at 752,6 size 35x35; Picture "ParlantesRojo"
      Visibility <- "SirenaChillers"
   Button "Botón_1" at 740,1 size 57x44; TextOff 'Text'
      on Click: ActivateScreen("MTA-ChillersConfiguraciónSirena", 0)
   TextField "Campo de texto_10" at 41,374 size 98x32; Text 'Presostato Agua Torres'
   Button "Botón_2" at 200,320 size 152x38; TextOff 'BOMBAS'
      on Click: ActivateScreen("MTA-TorreEnfriamientoBMB", 0)
   IOField "Campo ES_1" at 241,360 size 80x23; FormatPattern 999.99; Unit  ºC
      ProcessValue <- "TemperaturatorresCH"
   GraphicIOField "Campo ES gráfico_4" at 429,160 size 362x6; PictureList "Indicador"
      ProcessValue <- "AnimaciónV001"
   GraphicIOField "Campo ES gráfico_5" at 429,282 size 362x6; PictureList "Indicador"
      ProcessValue <- "AnimaciónV002"
   GraphicIOField "Campo ES gráfico_6" at 429,404 size 362x6; PictureList "Indicador"
      ProcessValue <- "AnimaciónV003"

Template "Plantilla_2" 800x480
   Button "Plantilla_1" at 640,429 size 78x48; TextOff 'Text'
   Button "Plantilla_8" at 81,429 size 78x48; TextOff 'Torres'
      on Release: ActivateScreen("MTA-TorreEnfriamientoBMB", 0)
   Button "Plantilla_10" at 2,429 size 78x48; TextOff 'Chillers'; TextOn 'NavigateHome'; PictureOff "NavigateHome_HMI_1"; PictureOn "NavigateHome_HMI_1"
      on Release: ActivateScreen("MTA-Chillers-General", 0)
   Button "Plantilla_11" at 720,429 size 78x48; TextOff 'Avisos'
      on Click: ActivateScreen("MTA-Avisos", 0)
      Appearance <- "AlarmaNueva"
   Button "Plantilla_2" at 480,429 size 78x48; TextOff 'Text'
   Button "Plantilla_3" at 560,429 size 78x48; TextOff 'Text'
   Button "Plantilla_4" at 400,429 size 78x48; TextOff 'Text'
   Button "Plantilla_5" at 320,429 size 78x48; TextOff 'Text'
   Button "Plantilla_6" at 240,429 size 78x48; TextOff 'Text'
   Button "Plantilla_7" at 160,429 size 78x48; TextOff 'Text'
   GraphicView "Plantilla_Visor de gráficos_26" at 68,9 size 91x26; Picture "eProC logo 4 b"
   GraphicView "Plantilla_Visor de gráficos_27" at 9,8 size 49x29; Picture "eProC logo 4 a"
*)

(* ===== HMI "HMI_RT_1" =====

text list "Enclavamientos": 0 'Ninguno'; 1 'ABC2'; 2 'ABC3'; 3 'Belliss'; 4 'ABC4'; 5 'ABC5'

ScreenModuleEditorView "Faceplate_7" 640x480
   GraphicView "Visor de gráficos_1" at 10,10 size 143x70; Picture "vlvV"
   GraphicView "Visor de gráficos_2" at 10,10 size 143x70; Picture "vlvR"
      Visibility <- "ON"
*)

(* ===== HMI "HMI_RT_1" =====
system functions are stored by id; their names below are inferred from use

text list "EstadoMotor": 0 'Detenido'; 1 'En Marcha'; 2 'Arrancando'; 3 'Deteniéndose'; 4 'Espera para Arrancar'; 5 'Sobrecarga de Corriente'; 6 'Deshabilitado'; 7 'En Falla'

ScreenModuleEditorView "ControlMotor-NoAUTO" 640x480
   Button "Botón_1" at 10,10 size 109x37; TextOff 'Habilitar'
      on Press: SetBit("Habilitación")
      on Release: ResetBit("Habilitación")
   Button "Botón_2" at 10,50 size 109x37; TextOff 'Deshabilitar'
      on Press: SetBit("Deshabilitación")
      on Release: ResetBit("Deshabilitación")
   Button "Botón_3" at 130,10 size 101x37; TextOff 'Marcha'
      on Press: SetBit("Marcha")
      on Release: ResetBit("Marcha")
   Button "Botón_4" at 130,50 size 101x37; TextOff 'Parada'
      on Press: SetBit("Parada")
      on Release: ResetBit("Parada")
*)

(* ===== HMI "HMI_RT_1" =====
system functions are stored by id; their names below are inferred from use

text list "Enclavamientos": 0 'Ninguno'; 1 'ABC2'; 2 'ABC3'; 3 'Belliss'; 4 'ABC4'; 5 'ABC5'

ScreenModuleEditorView "Faceplate_7" 640x480
   Button "Botón_3" at 25,15 size 189x37; TextOff 'Habilitar Marcha'
      on Press: SetBit("Marcha")
      Visibility <- "Animación"
      Appearance <- "Marcha"
   Button "Botón_1" at 11,10 size 93x40; TextOff 'MARCHA'
      on Press: SetBit("MARCHAF")
      Visibility <- "Animación"
      Appearance <- "MARCHAF"
   Button "Botón_2" at 11,54 size 93x40; TextOff 'PARADA'
      on Press: ResetBit("MARCHAF")
      Visibility <- "Animación"
      Appearance <- "MARCHAF"
   IOField "Campo ES_1" at 143,19 size 84x26; FormatPattern 999.99; Unit  bar
      ProcessValue <- "ON"
      Visibility <- "Animación"
   IOField "Campo ES_2" at 143,62 size 84x26; FormatPattern 999.99; Unit  bar
      ProcessValue <- "OFF"
      Visibility <- "Animación"
   TextField "Campo de texto_2" at 109,19 size 27x23; Text 'ON'
      Visibility <- "Animación"
   TextField "Campo de texto_3" at 109,62 size 32x23; Text 'OFF'
      Visibility <- "Animación"
   IOField "Campo ES_3" at 143,19 size 84x26; FormatPattern 999.99; Unit  bar
      ProcessValue <- "ON"
      Visibility <- "Animación"
   IOField "Campo ES_4" at 143,62 size 84x26; FormatPattern 999.99; Unit  bar
      ProcessValue <- "OFF"
      Visibility <- "Animación"
   TextField "Campo de texto_4" at 109,19 size 27x23; Text 'ON'
      Visibility <- "Animación"
   TextField "Campo de texto_5" at 109,62 size 32x23; Text 'OFF'
      Visibility <- "Animación"
   TextField "Campo de texto_1" at 10,31 size 97x40; Text 'Accionamiento Local'
      Visibility <- "Animación"
*)

(* ===== HMI "HMI_RT_1" =====
system functions are stored by id; their names below are inferred from use

text list "Enclavamientos": 0 'Ninguno'; 1 'ABC2'; 2 'ABC3'; 3 'Belliss'; 4 'ABC4'; 5 'ABC5'

ScreenModuleEditorView "Faceplate_2" 640x480
   TextField "Campo de texto_14" at 112,50 size 40x22; Text 'Enc 2'
      Visibility <- "Animación"
   TextField "Campo de texto_13" at 112,14 size 40x22; Text 'Enc 1'
      Visibility <- "Animación"
   Rectangle "Rectángulo_1" at 10,10 size 246x69
      Visibility <- "Animación"
   TextField "Campo de texto_1" at 67,18 size 125x50; Text 'Accionamiento Local'
      Visibility <- "Animación"
   Button "Botón_1" at 11,10 size 93x32; TextOff 'Habilitar'
      on Press: SetBit("Habilitación")
      on Release: ResetBit("Habilitación")
   Button "Botón_2" at 11,46 size 93x32; TextOff 'Deshabilitar'
      on Press: SetBit("Deshabilitación")
      on Release: ResetBit("Deshabilitación")
   Button "Botón_3" at 136,10 size 117x32; TextOff 'Marcha'
      on Press: SetBit("Marcha")
      on Release: ResetBit("Marcha")
      Visibility <- "Animación"
   Button "Botón_4" at 136,46 size 117x32; TextOff 'Parada'
      on Press: SetBit("Parada")
      on Release: ResetBit("Parada")
      Visibility <- "Animación"
   SymbolicIOField "Campo ES simbólico_2" at 158,12 size 96x27; TextOff '0'; TextOn '1'; TextList "Enclavamientos"
      ProcessValue <- "Enc1"
      Visibility <- "Animación"
   SymbolicIOField "Campo ES simbólico_3" at 158,47 size 96x27; TextOff '0'; TextOn '1'; TextList "Enclavamientos"
      ProcessValue <- "Enc2"
      Visibility <- "Animación"
*)

(* ===== HMI "HMI_RT_1" =====
system functions are stored by id; their names below are inferred from use

text list "EstadoMotor": 0 'Detenido'; 1 'En Marcha'; 2 'Arrancando'; 3 'Deteniéndose'; 4 'Espera para Arrancar'; 5 'Sobrecarga de Corriente'; 6 'Deshabilitado'; 7 'En Falla'

ScreenModuleEditorView "ControlMotor-NoAUTO" 640x480
   Button "Botón_1" at 10,10 size 109x37; TextOff 'Habilitar'
      on Press: SetBit("Habilitación")
      on Release: ResetBit("Habilitación")
   Button "Botón_2" at 10,50 size 109x37; TextOff 'Deshabilitar'
      on Press: SetBit("Deshabilitación")
      on Release: ResetBit("Deshabilitación")
   Button "Botón_3" at 130,10 size 101x37; TextOff 'Marcha'
      on Press: SetBit("Marcha")
      on Release: ResetBit("Marcha")
   Button "Botón_4" at 130,50 size 101x37; TextOff 'Parada'
      on Press: SetBit("Parada")
      on Release: ResetBit("Parada")
*)

(* ===== HMI "HMI_RT_1" =====
system functions are stored by id; their names below are inferred from use

ScreenModuleEditorView "Faceplate_4" 640x480
   TextField "Campo de texto_14" at 117,50 size 25x22; Text 'Off'
      Visibility <- "Animación"
   TextField "Campo de texto_13" at 119,14 size 23x22; Text 'On'
      Visibility <- "Animación"
   IOField "Campo ES_9" at 147,48 size 83x29; FormatPattern 999; Unit  ºC
      ProcessValue <- "SPOff"
      Visibility <- "Animación"
   IOField "Campo ES_8" at 147,12 size 83x29; FormatPattern 999; Unit  ºC
      ProcessValue <- "SPOn"
      Visibility <- "Animación"
   Button "Botón_1" at 10,10 size 93x32; TextOff 'Habilitar'
      on Press: SetBit("Habilitación")
      on Release: ResetBit("Habilitación")
   Button "Botón_2" at 10,46 size 93x32; TextOff 'Deshabilitar'
      on Press: SetBit("Deshabilitación")
      on Release: ResetBit("Deshabilitación")
   Button "Botón_3" at 122,10 size 109x32; TextOff 'Marcha'
      on Press: SetBit("Marcha")
      on Release: ResetBit("Marcha")
      Visibility <- "Animación"
   Button "Botón_4" at 122,46 size 109x32; TextOff 'Parada'
      on Press: SetBit("Parada")
      on Release: ResetBit("Parada")
      Visibility <- "Animación"
*)

(* ===== HMI "HMI_RT_1" =====
system functions are stored by id; their names below are inferred from use

ScreenModuleEditorView "Faceplate_1" 640x480
   TextField "Campo de texto_14" at 117,50 size 25x22; Text 'Off'
      Visibility <- "Animación"
   TextField "Campo de texto_13" at 119,14 size 23x22; Text 'On'
      Visibility <- "Animación"
   IOField "Campo ES_9" at 147,48 size 83x29; FormatPattern 999; Unit  ºC
      ProcessValue <- "SPOff"
      Visibility <- "Animación"
   IOField "Campo ES_8" at 147,12 size 83x29; FormatPattern 999; Unit  ºC
      ProcessValue <- "SPOn"
      Visibility <- "Animación"
   Button "Botón_1" at 10,10 size 93x32; TextOff 'Habilitar'
      on Press: SetBit("Habilitación")
      on Release: ResetBit("Habilitación")
   Button "Botón_2" at 10,46 size 93x32; TextOff 'Deshabilitar'
      on Press: SetBit("Deshabilitación")
      on Release: ResetBit("Deshabilitación")
   Button "Botón_3" at 122,10 size 109x32; TextOff 'Marcha'
      on Press: SetBit("Marcha")
      on Release: ResetBit("Marcha")
      Visibility <- "Animación"
   Button "Botón_4" at 122,46 size 109x32; TextOff 'Parada'
      on Press: SetBit("Parada")
      on Release: ResetBit("Parada")
      Visibility <- "Animación"
*)

(* ===== HMI "HMI_RT_1" =====
system functions are stored by id; their names below are inferred from use

ScreenModuleEditorView "Faceplate_1" 640x480
   TextField "Campo de texto_14" at 118,50 size 25x22; Text 'Off'
      Visibility <- "Animación"
   TextField "Campo de texto_13" at 120,14 size 23x22; Text 'On'
      Visibility <- "Animación"
   Rectangle "Rectángulo_1" at 10,10 size 227x69
      Visibility <- "Animación"
   TextField "Campo de texto_1" at 59,18 size 125x50; Text 'Accionamiento Local'
      Visibility <- "Animación"
   IOField "Campo ES_9" at 148,48 size 83x29; FormatPattern 99.99; Unit  bar
      ProcessValue <- "SPOff"
      Visibility <- "Animación"
   IOField "Campo ES_8" at 148,12 size 83x29; FormatPattern 99.99; Unit  bar
      ProcessValue <- "SPOn"
      Visibility <- "Animación"
   Button "Botón_1" at 11,10 size 93x32; TextOff 'Habilitar'
      on Press: SetBit("Habilitación")
      on Release: ResetBit("Habilitación")
   Button "Botón_2" at 11,46 size 93x32; TextOff 'Deshabilitar'
      on Press: SetBit("Deshabilitación")
      on Release: ResetBit("Deshabilitación")
   Button "Botón_3" at 123,10 size 109x32; TextOff 'Marcha'
      on Press: SetBit("Marcha")
      on Release: ResetBit("Marcha")
      Visibility <- "Animación"
   Button "Botón_4" at 123,46 size 109x32; TextOff 'Parada'
      on Press: SetBit("Parada")
      on Release: ResetBit("Parada")
      Visibility <- "Animación"
*)

(* ===== HMI "HMI_RT_1" =====
system functions are stored by id; their names below are inferred from use

text list "Enclavamientos": 0 'Ninguno'; 1 'ABC2'; 2 'ABC3'; 3 'Belliss'; 4 'ABC4'; 5 'ABC5'

ScreenModuleEditorView "Faceplate_10" 640x480
   Button "Botón_3" at 38,10 size 189x37; TextOff 'Habilitar Marcha'
      on Press: SetBit("Marcha")
      Visibility <- "Animación"
      Appearance <- "Marcha"
   Button "Botón_1" at 38,10 size 93x40; TextOff 'MARCHA'
      on Press: SetBit("MARCHAF")
      Visibility <- "Animación"
      Appearance <- "Forzando"
   Button "Botón_2" at 133,10 size 93x40; TextOff 'PARADA'
      on Press: ResetBit("MARCHAF")
      Visibility <- "Animación"
      Appearance <- "Forzando"
   IOField "Campo ES_1" at 44,75 size 84x26; FormatPattern 999.99; Unit  bar
      ProcessValue <- "ON"
      Visibility <- "Animación"
   IOField "Campo ES_2" at 44,110 size 84x26; FormatPattern 999.99; Unit  bar
      ProcessValue <- "OFF"
      Visibility <- "Animación"
   TextField "Campo de texto_2" at 10,75 size 27x23; Text 'ON'
      Visibility <- "Animación"
   TextField "Campo de texto_3" at 10,110 size 32x23; Text 'OFF'
      Visibility <- "Animación"
   IOField "Campo ES_3" at 140,75 size 84x26; FormatPattern 999.99; Unit  bar
      ProcessValue <- "ON2"
      Visibility <- "Animación"
   IOField "Campo ES_4" at 140,110 size 84x26; FormatPattern 999.99; Unit  bar
      ProcessValue <- "OFF2"
      Visibility <- "Animación"
   TextField "Campo de texto_4" at 60,51 size 45x23; Text 'Media'
      Visibility <- "Animación"
   TextField "Campo de texto_5" at 146,51 size 71x23; Text 'Completa'
      Visibility <- "Animación"
   IOField "Campo ES_5" at 44,75 size 84x26; FormatPattern 999.99; Unit  bar
      ProcessValue <- "ON"
      Visibility <- "Animación"
   IOField "Campo ES_6" at 44,110 size 84x26; FormatPattern 999.99; Unit  bar
      ProcessValue <- "OFF"
      Visibility <- "Animación"
   IOField "Campo ES_7" at 140,75 size 84x26; FormatPattern 999.99; Unit  bar
      ProcessValue <- "ON2"
      Visibility <- "Animación"
   IOField "Campo ES_8" at 140,110 size 84x26; FormatPattern 999.99; Unit  bar
      ProcessValue <- "OFF2"
      Visibility <- "Animación"
   TextField "Campo de texto_6" at 10,75 size 27x23; Text 'ON'
      Visibility <- "Animación"
   TextField "Campo de texto_7" at 10,110 size 32x23; Text 'OFF'
      Visibility <- "Animación"
   TextField "Campo de texto_8" at 60,51 size 45x23; Text 'Media'
      Visibility <- "Animación"
   TextField "Campo de texto_9" at 146,51 size 71x23; Text 'Completa'
      Visibility <- "Animación"
   TextField "Campo de texto_1" at 77,12 size 108x42; Text 'Accionamiento Local'
      Visibility <- "Animación"
*)

(* ===== HMI "HMI_RT_1" =====

ScreenModuleEditorView "Faceplate_6" 640x480
   GraphicIOField "PlotLight_Round_GN" at 52,10 size 35x34; PictureOff "PilotLight_Round_RN_Off_256c"; PictureOn "PilotLight_Round_GN_On_256c"
      ProcessValue <- "Verde"
      Visibility <- "Parpadeo"
   GraphicIOField "PlotLight_Round_RN" at 10,10 size 34x34; PictureOff "PilotLight_Round_RN_Off_256c"; PictureOn "PilotLight_Round_RN_On_256c"
      ProcessValue <- "Rojo"
   GraphicView "Visor de gráficos_1" at 52,10 size 34x34; Picture "PilotLight_Round_GN_Off_256c"
   GraphicView "Visor de gráficos_2" at 53,10 size 34x34; Picture "PilotLight_Round_GN_On_256c"
*)

(* ===== HMI "HMI_RT_1" =====
system functions are stored by id; their names below are inferred from use

ScreenModuleEditorView "Faceplate_1" 640x480
   Button "Botón_1" at 10,10 size 93x32; TextOff 'Habilitar'
      on Press: SetBit("Habilitación")
      on Release: ResetBit("Habilitación")
   Button "Botón_2" at 10,46 size 93x32; TextOff 'Deshabilitar'
      on Press: SetBit("Deshabilitación")
      on Release: ResetBit("Deshabilitación")
   Button "Botón_3" at 122,10 size 109x32; TextOff 'Marcha'
      on Press: SetBit("Marcha")
      on Release: ResetBit("Marcha")
   Button "Botón_4" at 122,46 size 109x32; TextOff 'Parada'
      on Press: SetBit("Parada")
      on Release: ResetBit("Parada")
*)

(* ===== HMI "HMI_RT_1" =====
system functions are stored by id; their names below are inferred from use
connection "Conexión-PLC_2": ETHERNET, SIMATIC S7 300/400 MPI
connection "Conexión-SentronPac_": ETHERNET, MODBUS_TCP

